(* Logix 5000 project; controller FV vendor 1 type 14 code 217 rev 31.11; software revision 31.00; part 15 of 63 *)
(* tags used below, declared in another part *)
   CWD : CHECKWORD_FLAGS;
   FR_AUDI1 : PlantItem;   // AUDI1
   FR_B246 : INT[255];   // V_REVERSE Flags for reversing contol action
   FR_BEACON1 : PlantItem;   // BEACON1
   FR_data_file_value_to_move : DINT;
   FR_F203 : REAL[40];
   FR_N100 : INT[265];   // FV FILLING
   FR_N110 : INT[265];   // GREEN BEER Green Beer Main
   FR_N120 : INT[265];   // YEAST CROP Yeast Cropping Main
   FR_N130 : INT[265];   // FILTRATE Filtrate Return
   FR_N14 : INT[265];   // MVFV CIP Comms to MVFV CIP Un it PLC
   FR_N140 : INT[265];   // CIP
   FR_N160 : INT[265];   // VESSEL Vessel Working Direc tory
   FR_N26 : INT[265];   // FV26
   FR_N27 : INT[265];   // FV27
   FR_N28 : INT[265];   // FV28
   FR_N29 : INT[265];   // FV29
   FR_N30 : INT[265];   // FV30
   FR_N31 : INT[265];   // FV31
   FR_N7 : INT[265];   // INTEGER
   FR_N99 : INT[265];   // COMMENT Comment Lines
   FR_PANELESTOP : PlantItem;   // PANELESTOP
   FR_PILZ : PlantItem;   // PILZ
   FR_T101 : TIMER[255];   // FV FILLING
   FR_T144 : TIMER[255];   // CIP
   FR_T4 : TIMER[255];   // TIMER
   FR_VB1_AV05 : PlantItem;   // VB1_AV05
   FR_VB1_AV08 : PlantItem;   // VB1_AV08
   FR_VB1_AV09 : PlantItem;   // VB1_AV09
   FR_VB2_AV01 : PlantItem;   // VB2_AV01
   FR_VB2_AV04 : PlantItem;   // VB2_AV04
   FR_VB2_AV05 : PlantItem;   // VB2_AV05
   FR_VB3_AV01 : PlantItem;   // VB3_AV01
   FR_VB3_AV04 : PlantItem;   // VB3_AV04
   FR_VB3_AV05 : PlantItem;   // VB3_AV05
(* FR_Common, continued *)

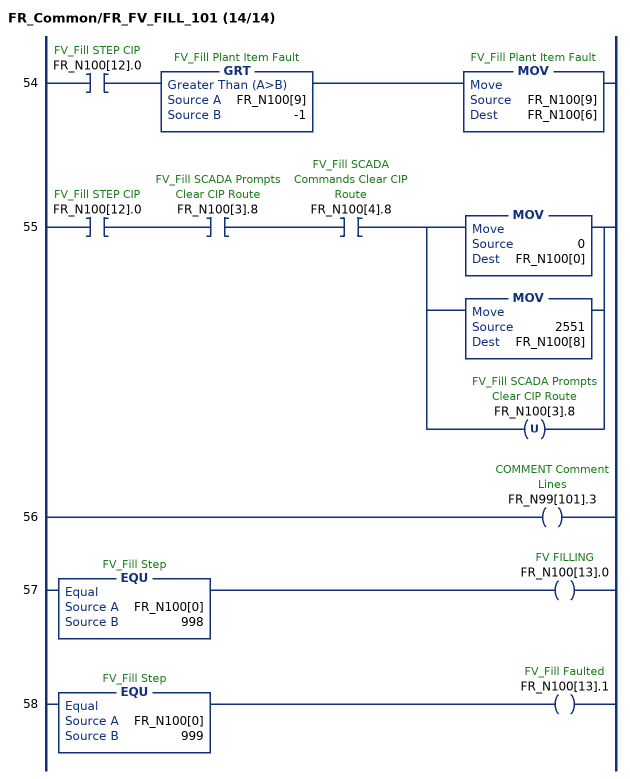
   [picture p230: FR_Common/FR_FV_FILL_101 rungs 54-58]
   54: XIC(FR_N100[12].0)GRT(FR_N100[9],-1)MOV(FR_N100[9],FR_N100[6]);
   55: XIC(FR_N100[12].0)XIC(FR_N100[3].8)XIC(FR_N100[4].8)[MOV(0,FR_N100[0]) ,MOV(2551,FR_N100[8]) ,OTU(FR_N100[3].8) ];
   56: OTE(FR_N99[101].3);
   57: EQU(FR_N100[0],998)OTE(FR_N100[13].0);
   58: EQU(FR_N100[0],999)OTE(FR_N100[13].1);
END_ROUTINE

ROUTINE FR_FV_FILL_OP_102   (* ladder *)
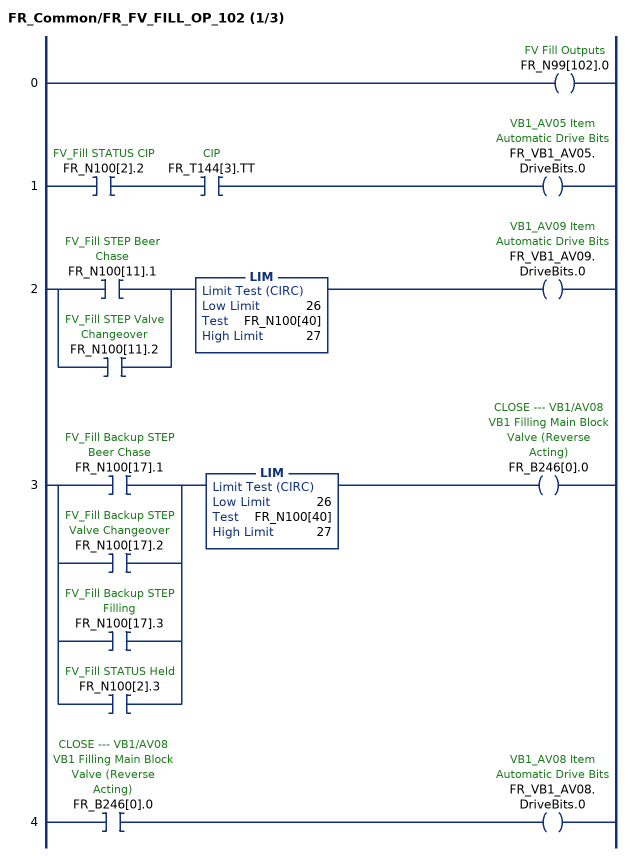
   0: OTE(FR_N99[102].0);
   1: XIC(FR_N100[2].2)XIC(FR_T144[3].TT)OTE(FR_VB1_AV05.DriveBits.0);
   2: [XIC(FR_N100[11].1) ,XIC(FR_N100[11].2) ]LIM(26,FR_N100[40],27)OTE(FR_VB1_AV09.DriveBits.0);
   3: [XIC(FR_N100[17].1) ,XIC(FR_N100[17].2) ,XIC(FR_N100[17].3) ,XIC(FR_N100[2].3) ]LIM(26,FR_N100[40],27)OTE(FR_B246[0].0);
   4: XIC(FR_B246[0].0)OTE(FR_VB1_AV08.DriveBits.0);
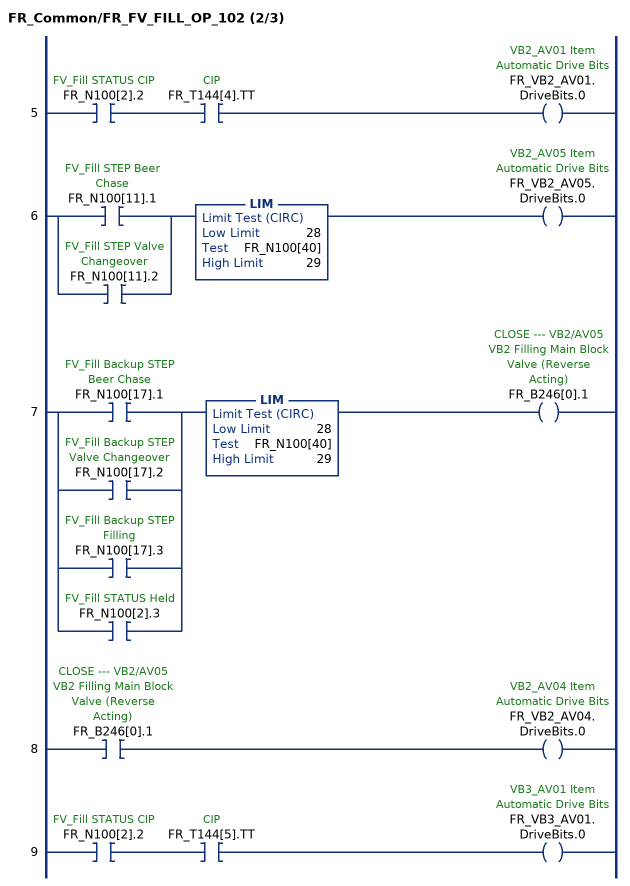
   5: XIC(FR_N100[2].2)XIC(FR_T144[4].TT)OTE(FR_VB2_AV01.DriveBits.0);
   6: [XIC(FR_N100[11].1) ,XIC(FR_N100[11].2) ]LIM(28,FR_N100[40],29)OTE(FR_VB2_AV05.DriveBits.0);
   7: [XIC(FR_N100[17].1) ,XIC(FR_N100[17].2) ,XIC(FR_N100[17].3) ,XIC(FR_N100[2].3) ]LIM(28,FR_N100[40],29)OTE(FR_B246[0].1);
   8: XIC(FR_B246[0].1)OTE(FR_VB2_AV04.DriveBits.0);
   9: XIC(FR_N100[2].2)XIC(FR_T144[5].TT)OTE(FR_VB3_AV01.DriveBits.0);
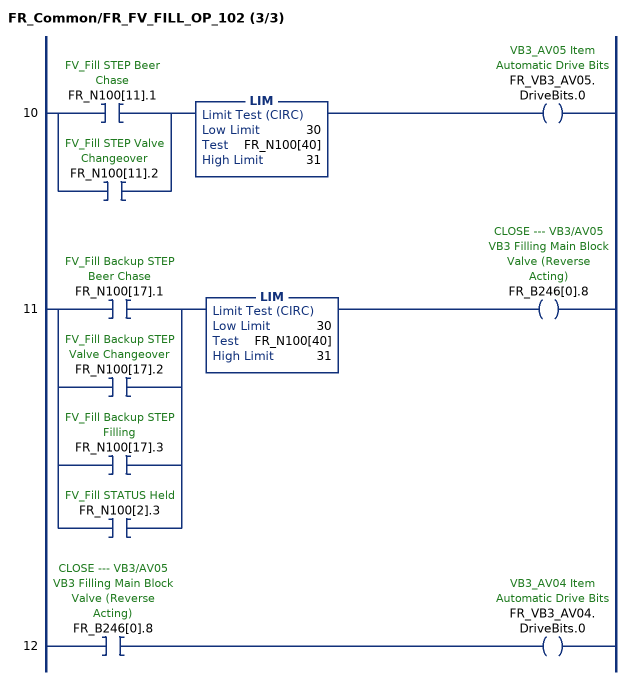
   10: [XIC(FR_N100[11].1) ,XIC(FR_N100[11].2) ]LIM(30,FR_N100[40],31)OTE(FR_VB3_AV05.DriveBits.0);
   11: [XIC(FR_N100[17].1) ,XIC(FR_N100[17].2) ,XIC(FR_N100[17].3) ,XIC(FR_N100[2].3) ]LIM(30,FR_N100[40],31)OTE(FR_B246[0].8);
   12: XIC(FR_B246[0].8)OTE(FR_VB3_AV04.DriveBits.0);
END_ROUTINE

ROUTINE FR_FV_FILL_ST_100   (* ladder *)
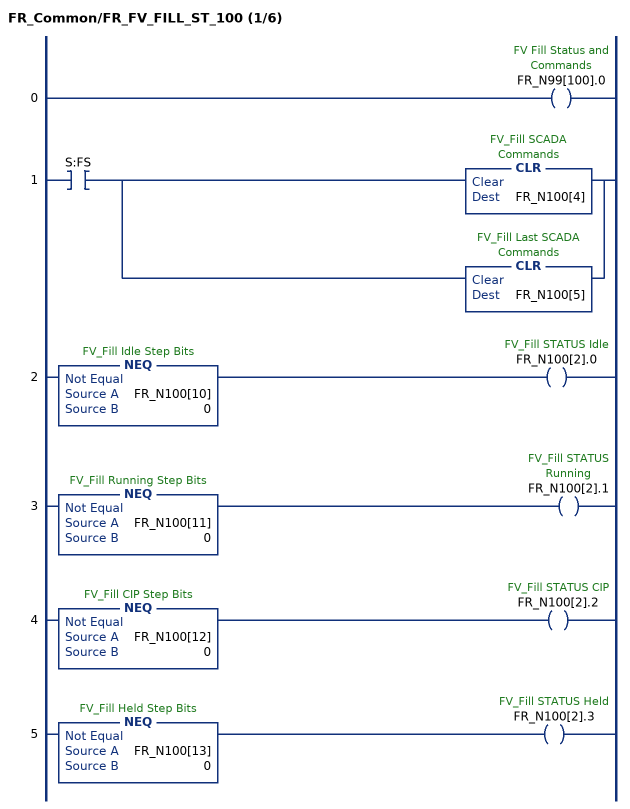
   0: OTE(FR_N99[100].0);
   1: XIC(S:FS)[CLR(FR_N100[4]) ,CLR(FR_N100[5]) ];
   2: NEQ(FR_N100[10],0)OTE(FR_N100[2].0);
   3: NEQ(FR_N100[11],0)OTE(FR_N100[2].1);
   4: NEQ(FR_N100[12],0)OTE(FR_N100[2].2);
   5: NEQ(FR_N100[13],0)OTE(FR_N100[2].3);
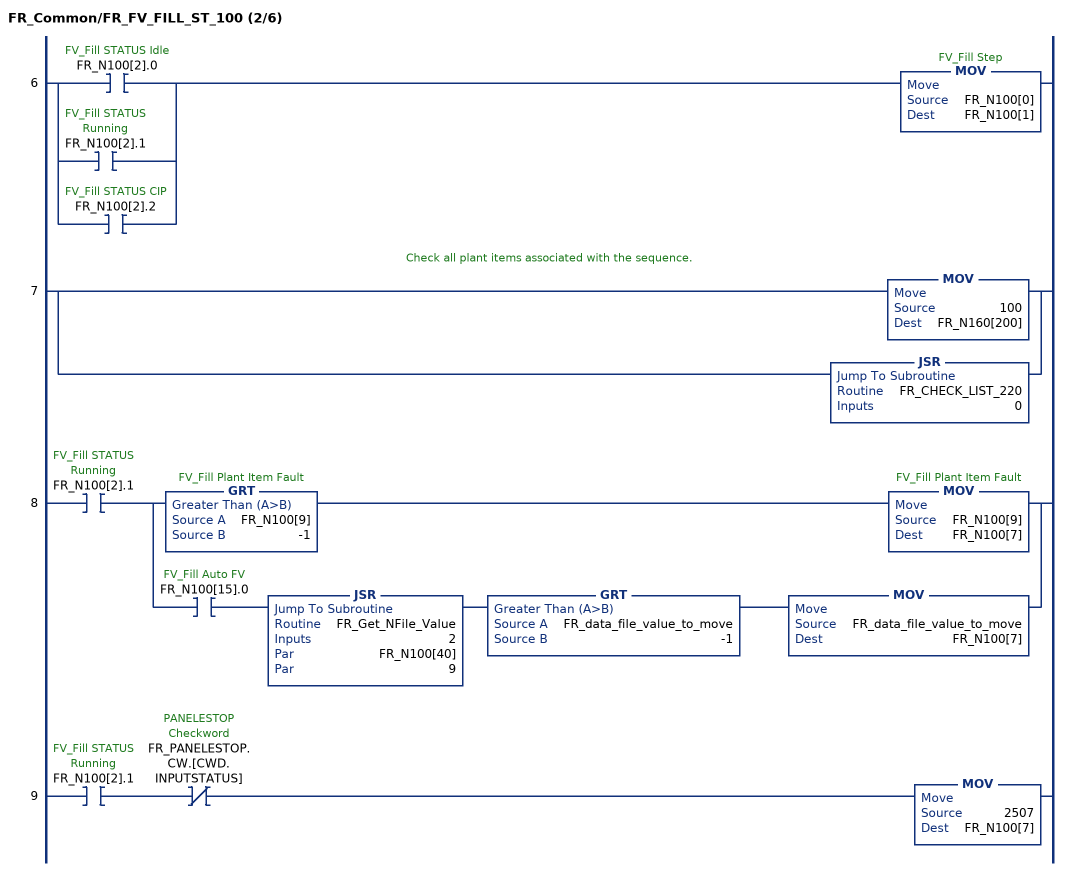
   6: [XIC(FR_N100[2].0) ,XIC(FR_N100[2].1) ,XIC(FR_N100[2].2) ]MOV(FR_N100[0],FR_N100[1]);
   // Check all plant items associated with the sequence.
   7: [MOV(100,FR_N160[200]) ,JSR(FR_CHECK_LIST_220,0) ];
   8: XIC(FR_N100[2].1)[GRT(FR_N100[9],-1) MOV(FR_N100[9],FR_N100[7]) ,XIC(FR_N100[15].0) JSR(FR_Get_NFile_Value,2,FR_N100[40],9) GRT(FR_data_file_value_to_move,-1) MOV(FR_data_file_value_to_move,FR_N100[7]) ];
   9: XIC(FR_N100[2].1)XIO(FR_PANELESTOP.CW.[CWD.INPUTSTATUS])MOV(2507,FR_N100[7]);
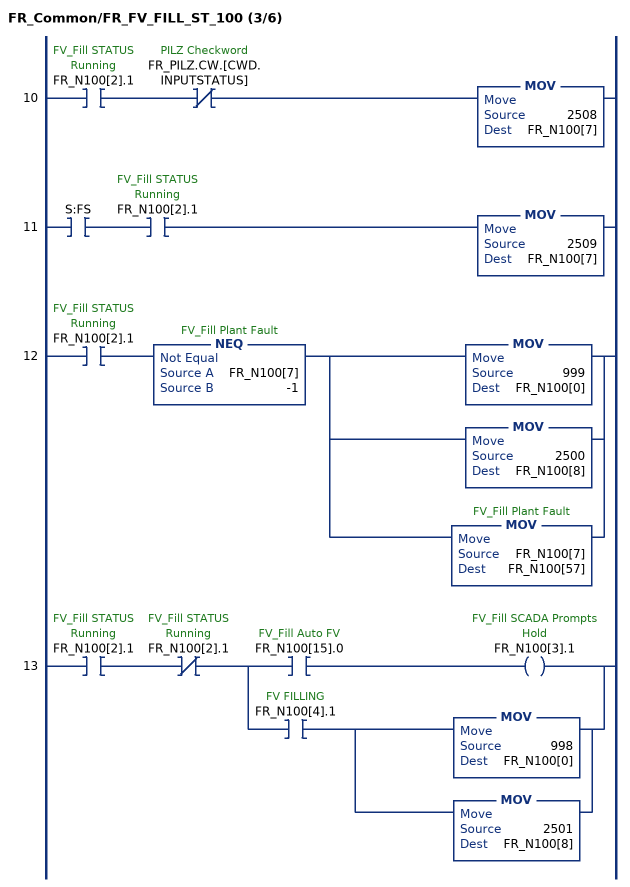
   10: XIC(FR_N100[2].1)XIO(FR_PILZ.CW.[CWD.INPUTSTATUS])MOV(2508,FR_N100[7]);
   11: XIC(S:FS)XIC(FR_N100[2].1)MOV(2509,FR_N100[7]);
   12: XIC(FR_N100[2].1)NEQ(FR_N100[7],-1)[MOV(999,FR_N100[0]) ,MOV(2500,FR_N100[8]) ,MOV(FR_N100[7],FR_N100[57]) ];
   13: XIC(FR_N100[2].1)XIO(FR_N100[2].1)[XIC(FR_N100[15].0) OTE(FR_N100[3].1) ,XIC(FR_N100[4].1) [MOV(998,FR_N100[0]) ,MOV(2501,FR_N100[8]) ] ];
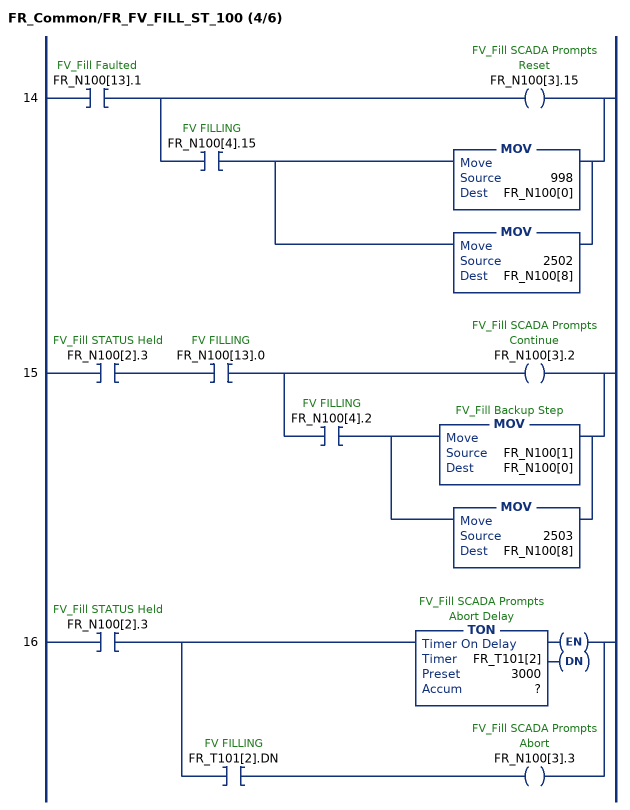
   14: XIC(FR_N100[13].1)[OTE(FR_N100[3].15) ,XIC(FR_N100[4].15) [MOV(998,FR_N100[0]) ,MOV(2502,FR_N100[8]) ] ];
   15: XIC(FR_N100[2].3)XIC(FR_N100[13].0)[OTE(FR_N100[3].2) ,XIC(FR_N100[4].2) [MOV(FR_N100[1],FR_N100[0]) ,MOV(2503,FR_N100[8]) ] ];
   16: XIC(FR_N100[2].3)[TON(FR_T101[2],?,?) ,XIC(FR_T101[2].DN) OTE(FR_N100[3].3) ];
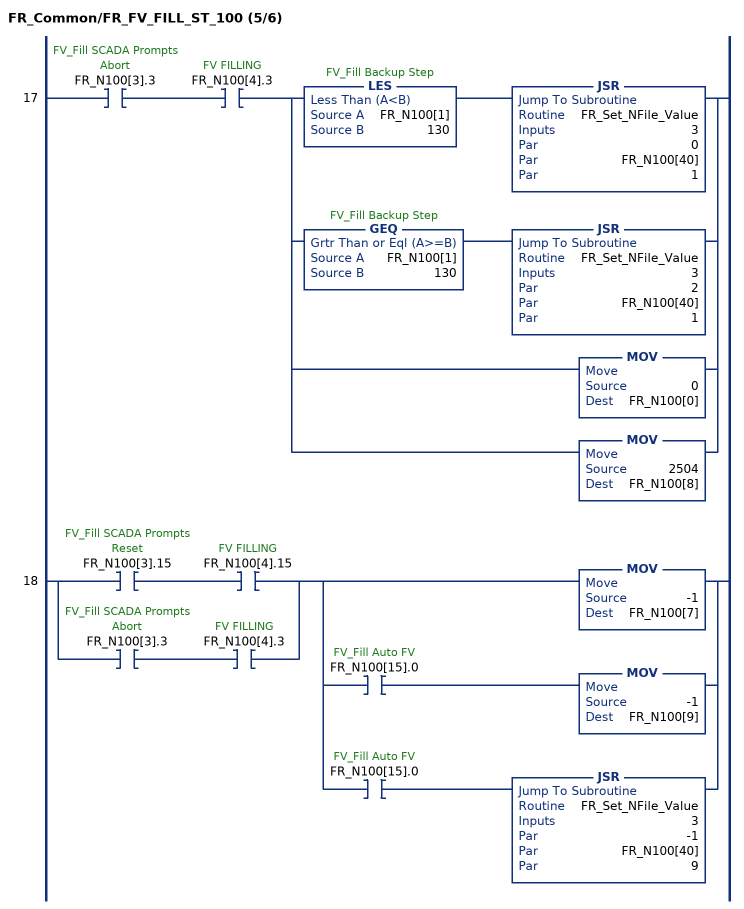
   17: XIC(FR_N100[3].3)XIC(FR_N100[4].3)[LES(FR_N100[1],130) JSR(FR_Set_NFile_Value,3,0,FR_N100[40],1) ,GEQ(FR_N100[1],130) JSR(FR_Set_NFile_Value,3,2,FR_N100[40],1) ,MOV(0,FR_N100[0]) ,MOV(2504,FR_N100[8]) ];
   18: [XIC(FR_N100[3].15) XIC(FR_N100[4].15) ,XIC(FR_N100[3].3) XIC(FR_N100[4].3) ][MOV(-1,FR_N100[7]) ,XIC(FR_N100[15].0) MOV(-1,FR_N100[9]) ,XIC(FR_N100[15].0) JSR(FR_Set_NFile_Value,3,-1,FR_N100[40],9) ];
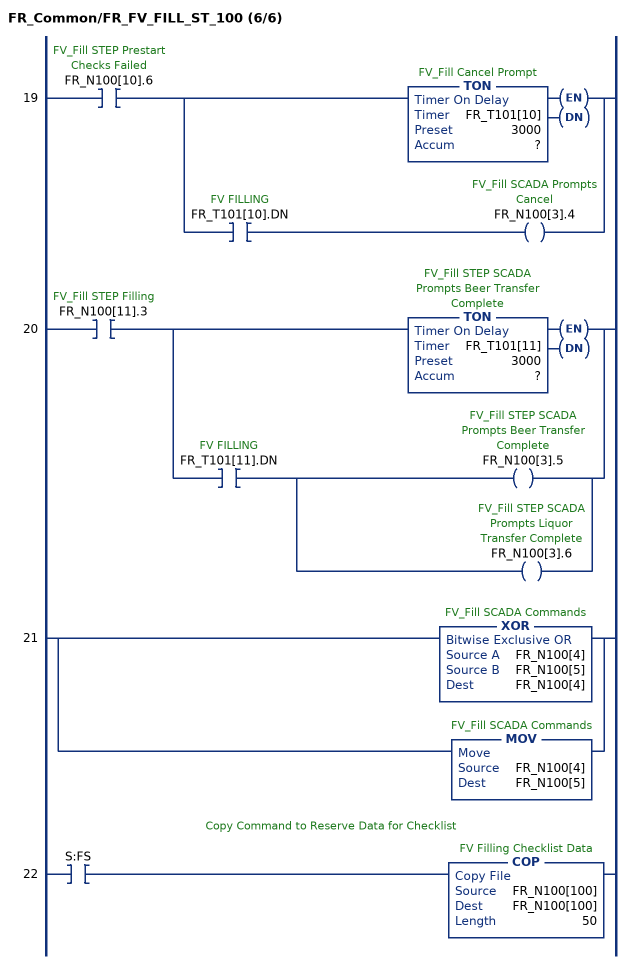
   19: XIC(FR_N100[10].6)[TON(FR_T101[10],?,?) ,XIC(FR_T101[10].DN) OTE(FR_N100[3].4) ];
   20: XIC(FR_N100[11].3)[TON(FR_T101[11],?,?) ,XIC(FR_T101[11].DN) [OTE(FR_N100[3].5) ,OTE(FR_N100[3].6) ] ];
   21: [XOR(FR_N100[4],FR_N100[5],FR_N100[4]) ,MOV(FR_N100[4],FR_N100[5]) ];
   // Copy Command to Reserve Data for Checklist
   22: XIC(S:FS)COP(FR_N100[100],FR_N100[100],50);
END_ROUTINE

ROUTINE FR_FV_VOLUME_202   (* ladder *)
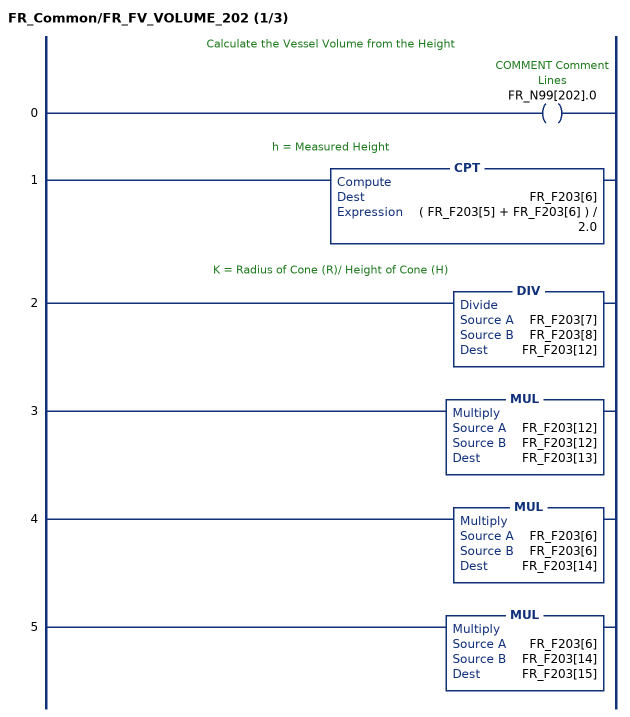
   // Calculate the Vessel Volume from the Height
   0: OTE(FR_N99[202].0);
   // h = Measured Height
   1: CPT(FR_F203[6],( FR_F203[5] + FR_F203[6] ) / 2.0);
   // K = Radius of Cone (R)/ Height of Cone (H)
   2: DIV(FR_F203[7],FR_F203[8],FR_F203[12]);
   3: MUL(FR_F203[12],FR_F203[12],FR_F203[13]);
   4: MUL(FR_F203[6],FR_F203[6],FR_F203[14]);
   5: MUL(FR_F203[6],FR_F203[14],FR_F203[15]);
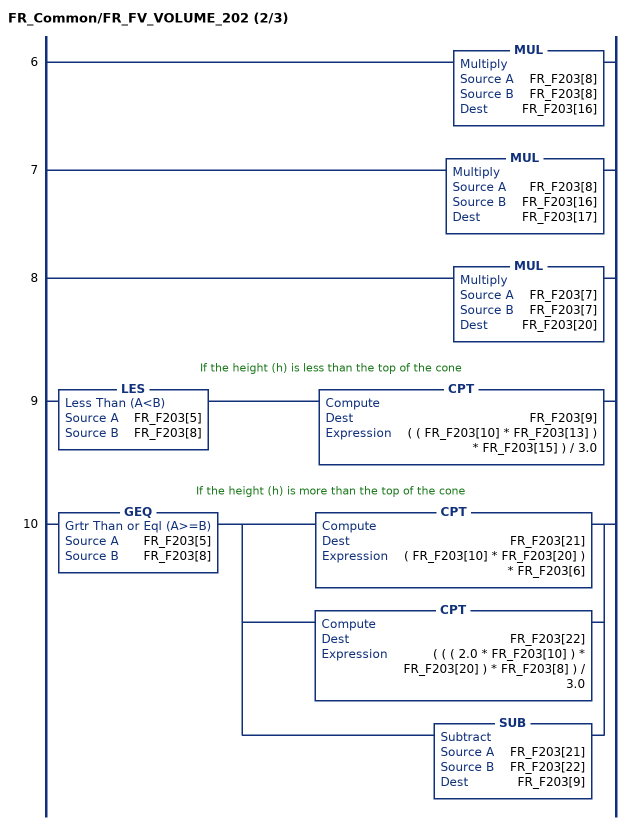
   6: MUL(FR_F203[8],FR_F203[8],FR_F203[16]);
   7: MUL(FR_F203[8],FR_F203[16],FR_F203[17]);
   8: MUL(FR_F203[7],FR_F203[7],FR_F203[20]);
   // If the height (h) is less than the top of the cone
   9: LES(FR_F203[5],FR_F203[8])CPT(FR_F203[9],( ( FR_F203[10] * FR_F203[13] ) * FR_F203[15] ) / 3.0);
   // If the height (h) is more than the top of the cone
   10: GEQ(FR_F203[5],FR_F203[8])[CPT(FR_F203[21],( FR_F203[10] * FR_F203[20] ) * FR_F203[6]) ,CPT(FR_F203[22],( ( ( 2.0 * FR_F203[10] ) * FR_F203[20] ) * FR_F203[8] ) / 3.0) ,SUB(FR_F203[21],FR_F203[22],FR_F203[9]) ];
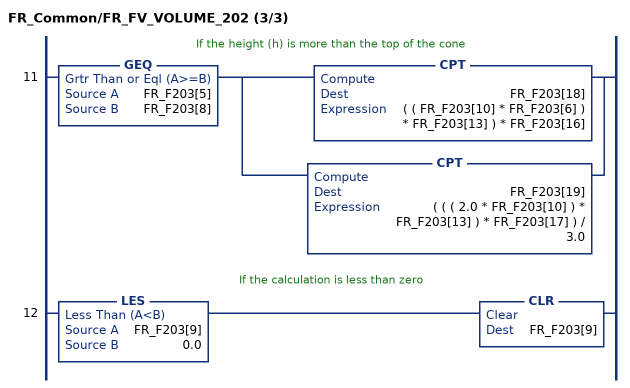
   // If the height (h) is more than the top of the cone
   11: GEQ(FR_F203[5],FR_F203[8])[CPT(FR_F203[18],( ( FR_F203[10] * FR_F203[6] ) * FR_F203[13] ) * FR_F203[16]) ,CPT(FR_F203[19],( ( ( 2.0 * FR_F203[10] ) * FR_F203[13] ) * FR_F203[17] ) / 3.0) ];
   // If the calculation is less than zero
   12: LES(FR_F203[9],0.0)CLR(FR_F203[9]);
END_ROUTINE

ROUTINE FR_GENERAL_7   (* ladder *)
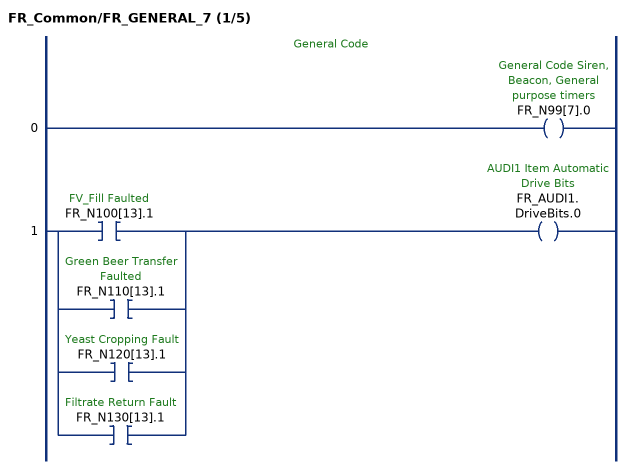
   // General Code
   0: OTE(FR_N99[7].0);
   1: [XIC(FR_N100[13].1) ,XIC(FR_N110[13].1) ,XIC(FR_N120[13].1) ,XIC(FR_N130[13].1) ]OTE(FR_AUDI1.DriveBits.0);
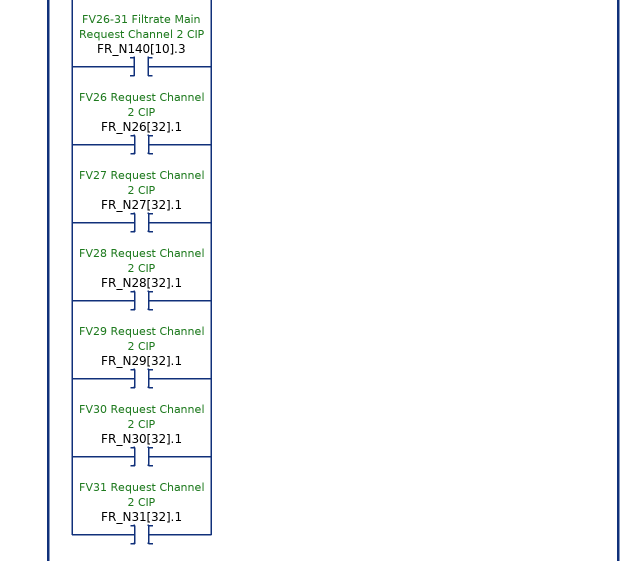
   2: [[XIC(FR_N140[0].0) ,XIC(FR_N140[0].1) ,XIC(FR_N140[0].2) ,XIC(FR_N140[0].3) ,XIC(FR_N26[32].0) ,XIC(FR_N27[32].0) ,XIC(FR_N28[32].0) ,XIC(FR_N29[32].0) ,XIC(FR_N30[32].0) ,XIC(FR_N31[32].0) ] XIC(FR_N14[4].5) ,[XIC(FR_N140[10].0) ,XIC(FR_N140[10].1) ,XIC(FR_N140[10].2) ,XIC(FR_N140[10].3) ,XIC(FR_N26[32].1) ,XIC(FR_N27[32].1) ,XIC(FR_N28[32].1) ,XIC(FR_N29[32].1) ,XIC(FR_N30[32].1) ,XIC(FR_N31[32].1) ] XIC(FR_N14[14].5) ]OTE(FR_BEACON1.DriveBits.0);
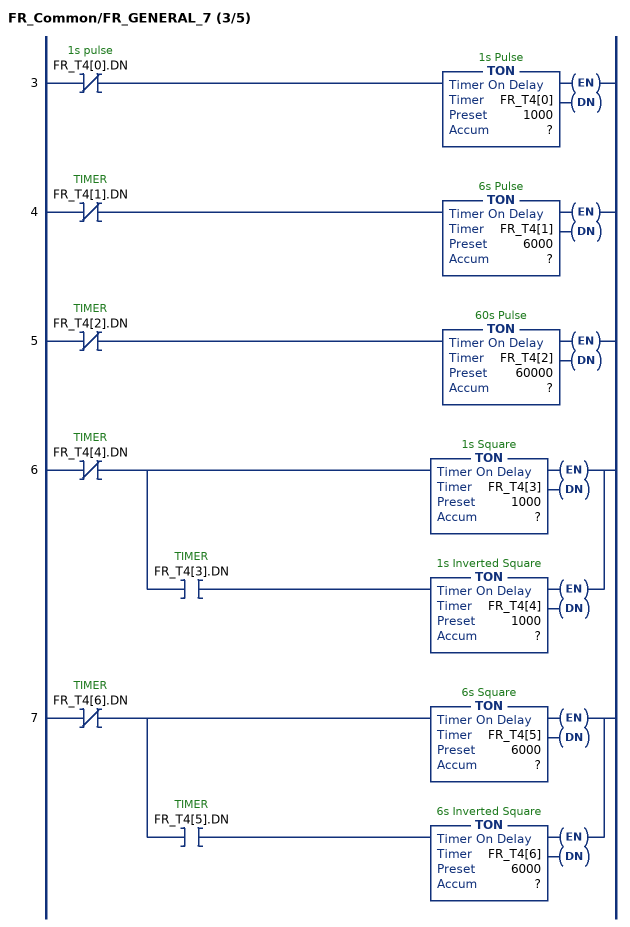
   3: XIO(FR_T4[0].DN)TON(FR_T4[0],?,?);
   4: XIO(FR_T4[1].DN)TON(FR_T4[1],?,?);
   5: XIO(FR_T4[2].DN)TON(FR_T4[2],?,?);
   6: XIO(FR_T4[4].DN)[TON(FR_T4[3],?,?) ,XIC(FR_T4[3].DN) TON(FR_T4[4],?,?) ];
   7: XIO(FR_T4[6].DN)[TON(FR_T4[5],?,?) ,XIC(FR_T4[5].DN) TON(FR_T4[6],?,?) ];
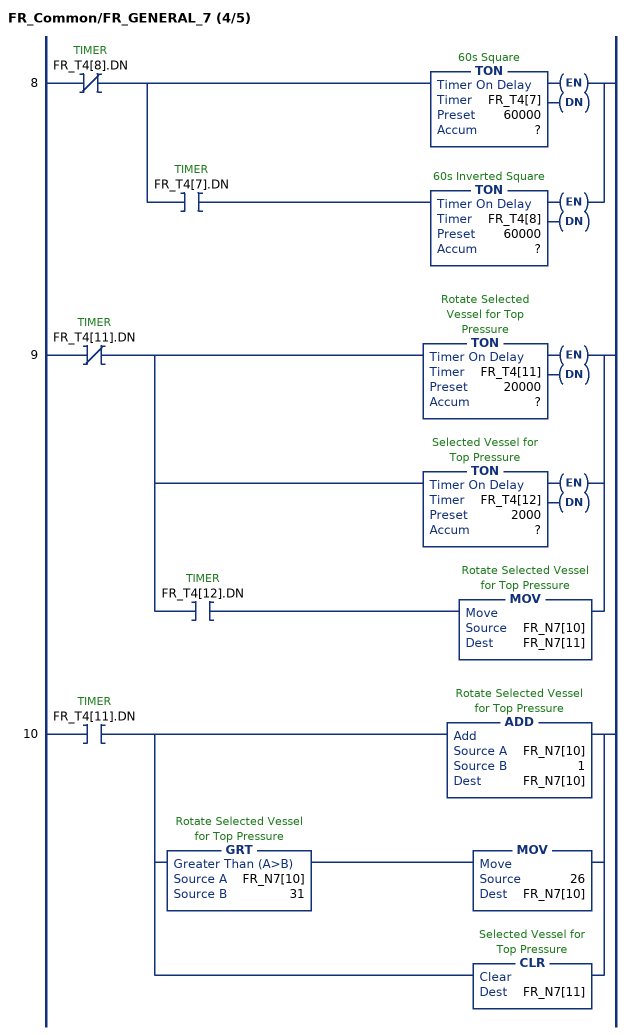
   8: XIO(FR_T4[8].DN)[TON(FR_T4[7],?,?) ,XIC(FR_T4[7].DN) TON(FR_T4[8],?,?) ];
   9: XIO(FR_T4[11].DN)[TON(FR_T4[11],?,?) ,TON(FR_T4[12],?,?) ,XIC(FR_T4[12].DN) MOV(FR_N7[10],FR_N7[11]) ];
   10: XIC(FR_T4[11].DN)[ADD(FR_N7[10],1,FR_N7[10]) ,GRT(FR_N7[10],31) MOV(26,FR_N7[10]) ,CLR(FR_N7[11]) ];
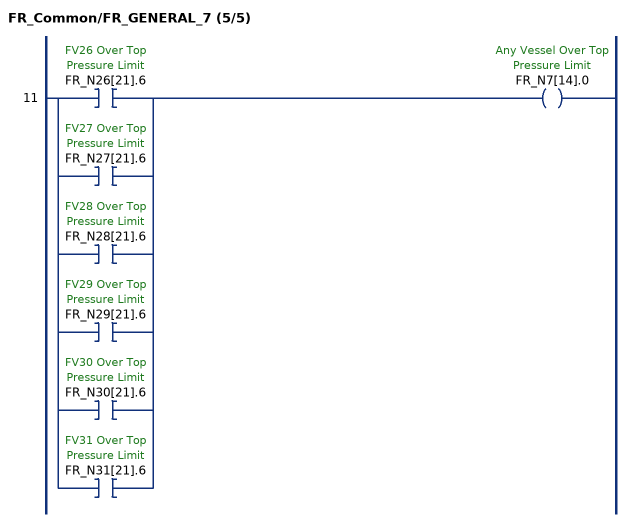
   11: [XIC(FR_N26[21].6) ,XIC(FR_N27[21].6) ,XIC(FR_N28[21].6) ,XIC(FR_N29[21].6) ,XIC(FR_N30[21].6) ,XIC(FR_N31[21].6) ]OTE(FR_N7[14].0);
END_ROUTINE
